// TIA Portal project "EdgeHowTos" (V16)

(* hardware
DEVICE "S71500/ET200MP station_1"  S7-1500 station
   slot 0: "Rail_0"  Rack  6ES7 590-1***0-0AA0
   slot 1: "PLC"  CPU 1513-1 PN  6ES7 513-1AL02-0AB0  V2.8
      slot 3: "CPU display_1"  6ES7591-1AA00-0AA0
      slot 32768: "PROFINET interface_1"  X1
         slot 32769: "Port_1"  X1 P1
         slot 32770: "Port_2"  X1 P2
      slot 34817: "Virtual CP interface port_1"  Virtual CP interface port  Virtual CP interface port
DEVICE "HMI"  TP900 Comfort
   slot 0: "HMI"  TP900 Comfort  6AV2 124-0JC01-0AX0  16.0.0.0
   slot 1: "HMI_RT_5"  TP900 Comfort  6AV2 124-0JC01-0AX0  16.0.0.0
   slot 5: "HMI._CP_1"  PROFINET Interface  16.0.0.0
      slot 1: "PROFINET Interface_1"  PROFINET Interface
         slot 1: "Port_1"  Port
         slot 2: "Port_2"  Port
   slot 7: "HMI.I/DP_CP_1"  MPI/DP Interface  16.0.0.0
*)

// ===== PLC "PLC"  CPU 1513-1 PN =====

VAR_GLOBAL   // PLC tag table "Default tag table"
   "Manipulator" AT %MW0 : Int;
END_VAR

VAR_GLOBAL CONSTANT   // PLC tag table "Default tag table"
   "STATE_FILL_TANK" : Int := 1;
   "STATE_HEAT_TANK" : Int := 2;
   "STATE_FILL_BOTTLE" : Int := 3;
   "STATE_SHIFT_BOTTLE" : Int := 4;
   "STATE_STOP" : Int := 5;
   "STATE_RESET" : Int := 6;
   "STATE_ERROR" : Int := 7;
   "ERROR_0_NO" : UInt := 0;
   "ERROR_1_CONNECTION" : UInt := 1;
   "ERROR_2_POWER" : UInt := 2;
   "ERROR_3_MANPOWER" : UInt := 3;
   "ERROR_4_CONVEYOR" : UInt := 4;
   "ERROR_5_VENTIL" : UInt := 5;
   "ERROR_6_HEATING" : UInt := 6;
   "ERROR_7_BOTTLE" : UInt := 7;
END_VAR

TYPE "typeHmi"
   STRUCT
      HMI_Start : Bool;   // trigger from hmi to start
      HMI_Stop : Bool;   // trigger from hmi to stop
      HMI_Reset : Bool;   // trigger from hmi to reset
      HMI_NextBottle : Bool;   // trigger from hmi to shift bottle
      HMI_Error : Bool;   // trigger from hmi to generate error
   END_STRUCT;
END_TYPE

TYPE "typeApp"
   STRUCT
      APP_Start : Bool;   // trigger from app to start
      APP_Stop : Bool;   // trigger from app to stop
      APP_Reset : Bool;   // trigger from app to reset
      APP_QRCode : String;   // string from app containing QR code (scanning app)
      APP_NextBottle : Bool;   // trigger from app to shift bottle
      APP_Error : Bool;   // trigger from app to generate error
      APP_Alarm : Bool;   // trigger from app to generate program alarm
   END_STRUCT;
END_TYPE

TYPE "typeSignals"
   STRUCT
      tankSignals : Struct
         actLevel : Real;   // actual level of tank [l]
         maxLevel : Bool;   // max level of tank reached
         actPressure : Real;   // actual pressure of tank [hPa]
         actTemperature : Real;   // actual temperature of tank [°C]
         maxTemperature : Bool;   // max level of temperature reached
      END_STRUCT;
      bottleSignals : Struct
         actLevel : Real;   // actual level of current bottle [l]
         maxLevel : Bool;   // max level of bottle reached
         outputTank : Real;   // Vout of Tank / Vin of bottle [m³/s]
      END_STRUCT;
      energySignals : Struct
         energyConsumptionFillingTank : Real;   // energy consumption during filling tank [Wh]
         waterConsumptionFillingTank : Real;   // water consumption during filling tank [l]
         energyConsumptionHeatingTank : Real;   // energy consumption during heating tank [Wh]
         energyConsumptionFillingBottles : Real;   // energy consumption during filling bottles [Wh]
         gasConsumptionHeatingTank : Real;   // gas consumption during heating tank [Wh]
      END_STRUCT;
      alarm : Word;   // alarm bit
   END_STRUCT;
END_TYPE

TYPE "typeOperate"
   STRUCT
      extModeActive : Bool := false;   // true = activate external model / simulation
      state : "typeState";   // operating state
      machineState : Int := 0;   // see user constants (1 = filling tank, 2 = heating tank, 3 = filling bottle, 4 = shifting bottle, 5 = stop, 6 = reset)
   END_STRUCT;
END_TYPE

TYPE "typeModel"
   STRUCT
      cycleTime : Real;   // cycle time[s]
      tank : Struct   // model struct of tank
         AT : Real;   // surface area of tank [m²]
         H : Real;   // high of tank [m]
         Vin : Real;   // incoming volume flow [l/min]
         maxLevel : Real;   // max level of tank [m³]
         roomTemperature : Real;   // room temperature of tank [°C]
         maxTemperature : Real;   // max temperature of tank [°C]
         density : Real;   // liquid density [kg/m³]
      END_STRUCT;
      bottle : Struct   // model struct of bottle
         maxLevel : Real;   // max level of bottle [m³]
         AB : Real;   // surface area of filling hole to fill bottle [m²]
      END_STRUCT;
   END_STRUCT;
END_TYPE

TYPE "typeProcess"
   STRUCT
      productId : UDInt;   // product id of current bottle
      numberProduced : UDInt;   // number of filled bottles
      numberFaulty : UDInt;   // number of faulty bottles
      batchId : UDInt;   // batch id (according to tank filling)
   END_STRUCT;
END_TYPE

TYPE "typeState"
   STRUCT
      FillingTank : Bool;   // filling tank
      HeatingTank : Bool;   // heating tank
      FillingBottle : Bool;   // filling bottle
      ShiftingBottle : Bool;   // shifting bottle
      Stop : Bool;   // stop filling application
      Reset : Bool;   // reset application
      Error : Bool;   // error within filling application
   END_STRUCT;
END_TYPE

TYPE "typeInfo"
   STRUCT
      "version" : String;   // current version of the project
      "date" : String;   // last change date of the project
   END_STRUCT;
END_TYPE

TYPE "typeError"
   STRUCT
      errorSimulation : Bool := true;   // activate simulation
      errorTrigger : Bool := false;   // trigger manual error simulation
      errorDuration : Time := T#120s;   // error duration for simlation
      errorCode : UInt := 0;   // error code for error analysis
   END_STRUCT;
END_TYPE

DATA_BLOCK "GDB"   // DB1
{ S7_Optimized_Access := 'FALSE' }
VERSION : 0.1
   VAR
      operate : "typeOperate";   // application operation
      model : "typeModel";   // model parameter
      externalSignals : "typeSignals";   // signals from external model
      signals : "typeSignals";   // current signals from tank and bottle
      process : "typeProcess";   // current process information
      hmiSignals : "typeHmi";   // signals from hmi
      appSignals : "typeApp";   // signals from edge app
      projectInfo : "typeInfo";   // infos regarding this TIA project
      errors : "typeError";
   END_VAR
BEGIN
   model.tank.H := 2.0;
   model.tank.AT := 0.8;
   operate.extModeActive := false;
   model.tank.maxTemperature := 80.0;
   model.tank.maxLevel := 1.6;
   model.bottle.maxLevel := 0.1;
   model.cycleTime := 0.01;
   model.tank.roomTemperature := 20.0;
   model.tank.Vin := 500.0;
   model.bottle.AB := 0.001;
   process.productId := 0;
   process.numberProduced := 0;
   process.numberFaulty := 0;
   model.tank.density := 997.0;
   hmiSignals.HMI_Start := true;
   projectInfo."version" := 'V1.1';
   projectInfo."date" := '2024-04-18';
END_DATA_BLOCK

DATA_BLOCK "DB_1_Sequence"   // DB2
{ S7_Optimized_Access := 'TRUE' }
VERSION : 0.1
// stored: InstanceOfName FB_1_Sequence
"FB_1_Sequence"
BEGIN
END_DATA_BLOCK

DATA_BLOCK "DB_2_Filling_DB"   // DB3
{ S7_Optimized_Access := 'TRUE' }
VERSION : 0.1
// stored: InstanceOfName FB_2_Filling
"FB_2_Filling"
BEGIN
END_DATA_BLOCK

DATA_BLOCK "DB_3_Simulation"   // DB4
{ S7_Optimized_Access := 'TRUE' }
VERSION : 0.1
// stored: InstanceOfName FB_3_Simulation
"FB_3_Simulation"
BEGIN
END_DATA_BLOCK

FUNCTION_BLOCK "FB_1_Sequence"   // FB2, FBD
{ S7_Optimized_Access := 'TRUE' }
VERSION : 0.1
   VAR_INPUT
      model : "typeModel";   // model parameter
      externalSignals : "typeSignals";   // signals from external model
   END_VAR
   VAR_IN_OUT
      operate : "typeOperate";   // application operation
      signals : "typeSignals";   // current signals from tank
      process : "typeProcess";   // current process information
      hmi : "typeHmi";   // signals from hmi
      app : "typeApp";   // signals from app
      errors : "typeError";
   END_VAR
   VAR
      statStart : Bool;   // trigger for start command
      statStop : Bool;   // trigger for stop command
      statReset : Bool;   // trigger for reset command
      statInit : Bool := true;   // helper variable to initialize some parameters
      statNextBottle : Bool;   // trigger to shift next bottle
      statError : Bool;   // trigger to set error
      statState : Int;   // memory for reactivating state after STOP
      statAlarm : Bool;   // trigger to generate program alarm
      statMemoryStart : Bool;
      statMemoryStop : Bool;
      statMemoryReset : Bool;
      statMemoryNextBottle : Bool;
      statMemoryError : Bool;
      statHmiStateStart : Bool;   // helper for hmi (true, if state 1-4)
      statShiftingTimer : Int;
      statShiftingTimerTrigger : Bool;
      statShiftingTrigger : Bool;
      statShiftingTimerDone : Bool;
      statHmiQrCodeReceived : Bool;
      statHMIQrCodeReceivedTrigger : Bool;
      statQrCodeTrigger : Bool;
      statTankEmpty : Bool;   // trigger when tank is empty
      statTankEmptyMemory : Bool;   // tank empty memory
      statOverflow : Bool;   // overflow of counter "numberProduced"
      statOverflowStartTrigger : Bool;   // trigger to start after overflow
      statOverflowStartMemory : Bool;
      Program_Alarm : Program_Alarm;
   END_VAR
   VAR_TEMP
      tempQrCodeLen : Int;
      tempProgramAlarmError : Bool;
      tempProgramAlarmStatus : Word;
      tempAlarmStateError : Bool;
      tempAlarmStateStatus : Word;
   END_VAR
   VAR_TEMP   // added for the SCL form of the ladder/FBD networks
      _w1 : Bool;
      _w2 : Bool;
      _w3 : Bool;
      _w4 : Bool;
   END_VAR
BEGIN

REGION Network 1: Handling signals from hmi or app
   // --[P]-- (positive signal edge) -> stat-Variable becomes true for one cycle
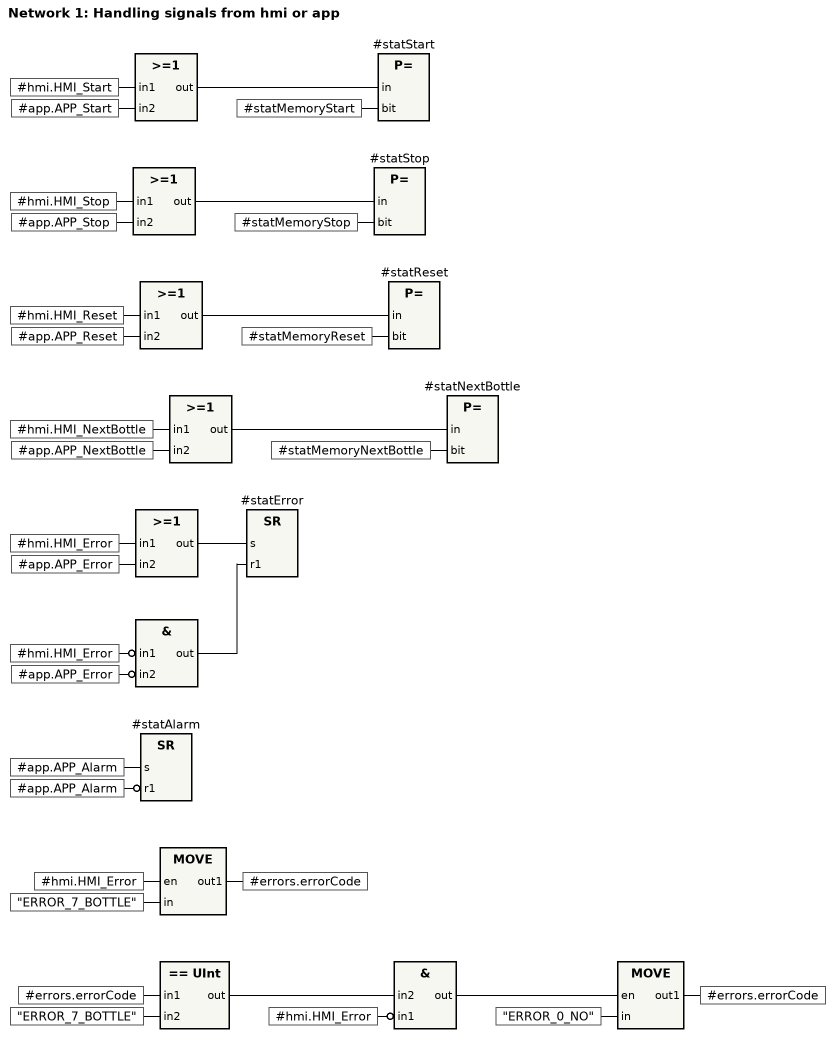
   #_w1 := #hmi.HMI_Start OR #app.APP_Start;
   #statStart := #_w1 AND NOT #statMemoryStart;   // rising edge
   #statMemoryStart := #_w1;
   #_w2 := #hmi.HMI_Stop OR #app.APP_Stop;
   #statStop := #_w2 AND NOT #statMemoryStop;   // rising edge
   #statMemoryStop := #_w2;
   #_w3 := #hmi.HMI_Reset OR #app.APP_Reset;
   #statReset := #_w3 AND NOT #statMemoryReset;   // rising edge
   #statMemoryReset := #_w3;
   #_w4 := #hmi.HMI_NextBottle OR #app.APP_NextBottle;
   #statNextBottle := #_w4 AND NOT #statMemoryNextBottle;   // rising edge
   #statMemoryNextBottle := #_w4;
   IF #hmi.HMI_Error OR #app.APP_Error THEN
       #statError := TRUE;   // SR flip-flop
   END_IF;
   IF NOT #hmi.HMI_Error AND NOT #app.APP_Error THEN #statError := FALSE; END_IF;
   IF #app.APP_Alarm THEN
       #statAlarm := TRUE;   // SR flip-flop
   END_IF;
   IF NOT #app.APP_Alarm THEN #statAlarm := FALSE; END_IF;
   IF #hmi.HMI_Error THEN #errors.errorCode := "ERROR_7_BOTTLE"; END_IF;
   IF (#errors.errorCode = "ERROR_7_BOTTLE") AND NOT #hmi.HMI_Error THEN
       #errors.errorCode := "ERROR_0_NO";
   END_IF;
END_REGION

REGION Network 2: Reset signals from hmi or app
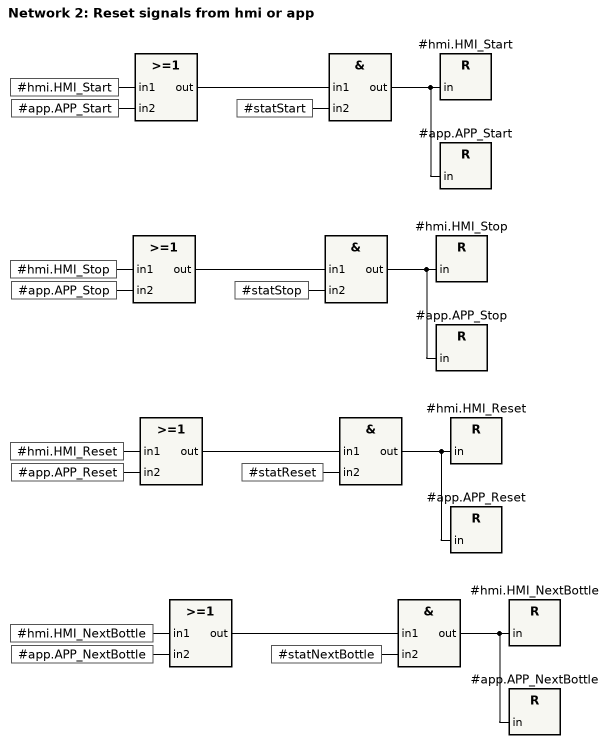
   #_w1 := (#hmi.HMI_Start OR #app.APP_Start) AND #statStart;
   IF #_w1 THEN
       #hmi.HMI_Start := FALSE;
       #app.APP_Start := FALSE;
   END_IF;
   #_w2 := (#hmi.HMI_Stop OR #app.APP_Stop) AND #statStop;
   IF #_w2 THEN
       #hmi.HMI_Stop := FALSE;
       #app.APP_Stop := FALSE;
   END_IF;
   #_w3 := (#hmi.HMI_Reset OR #app.APP_Reset) AND #statReset;
   IF #_w3 THEN
       #hmi.HMI_Reset := FALSE;
       #app.APP_Reset := FALSE;
   END_IF;
   #_w4 := (#hmi.HMI_NextBottle OR #app.APP_NextBottle) AND #statNextBottle;
   IF #_w4 THEN
       #hmi.HMI_NextBottle := FALSE;
       #app.APP_NextBottle := FALSE;
   END_IF;
END_REGION

REGION Network 3: Helper for hmi display
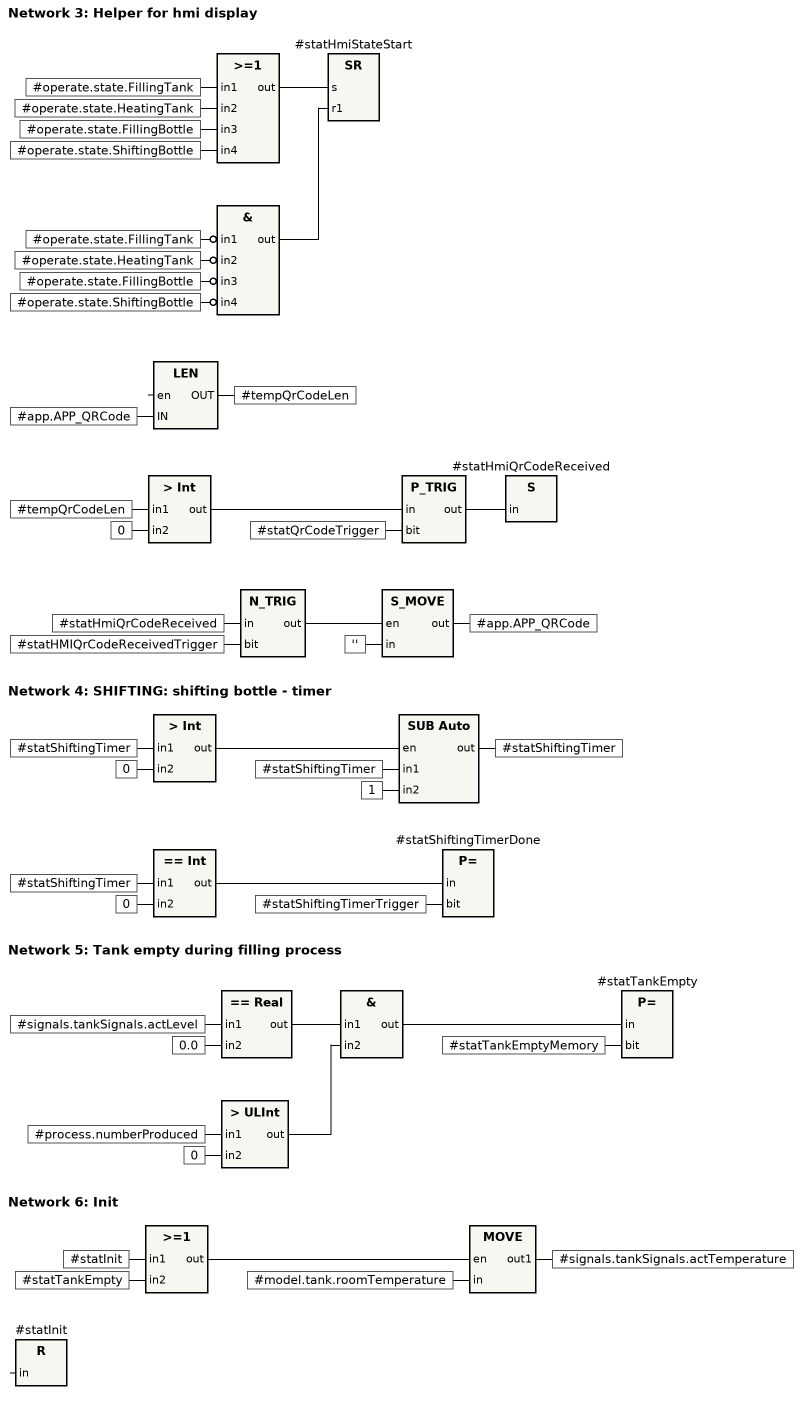
   IF #operate.state.FillingTank OR #operate.state.HeatingTank OR #operate.state.FillingBottle OR #operate.state.ShiftingBottle THEN
       #statHmiStateStart := TRUE;   // SR flip-flop
   END_IF;
   IF NOT #operate.state.FillingTank AND NOT #operate.state.HeatingTank AND NOT #operate.state.FillingBottle AND NOT #operate.state.ShiftingBottle THEN
       #statHmiStateStart := FALSE;
   END_IF;
   #tempQrCodeLen := LEN(IN := #app.APP_QRCode);
   #_w1 := #tempQrCodeLen > 0;
   #_w2 := #_w1 AND NOT #statQrCodeTrigger;   // rising edge
   #statQrCodeTrigger := #_w1;
   IF #_w2 THEN #statHmiQrCodeReceived := TRUE; END_IF;
   #_w3 := NOT #statHmiQrCodeReceived AND #statHMIQrCodeReceivedTrigger;   // falling edge
   #statHMIQrCodeReceivedTrigger := #statHmiQrCodeReceived;
   IF #_w3 THEN #app.APP_QRCode := ''; END_IF;
END_REGION

REGION Network 4: SHIFTING: shifting bottle - timer
   IF #statShiftingTimer > 0 THEN #statShiftingTimer := #statShiftingTimer - 1; END_IF;
   #_w1 := #statShiftingTimer = 0;
   #statShiftingTimerDone := #_w1 AND NOT #statShiftingTimerTrigger;   // rising edge
   #statShiftingTimerTrigger := #_w1;
END_REGION

REGION Network 5: Tank empty during filling process
   #_w1 := (#signals.tankSignals.actLevel = 0.0) AND (#process.numberProduced > 0);
   #statTankEmpty := #_w1 AND NOT #statTankEmptyMemory;   // rising edge
   #statTankEmptyMemory := #_w1;
END_REGION

REGION Network 6: Init
   IF #statInit OR #statTankEmpty THEN
       #signals.tankSignals.actTemperature := #model.tank.roomTemperature;
   END_IF;
   #statInit := FALSE;
END_REGION

REGION Network 7: Filling tank
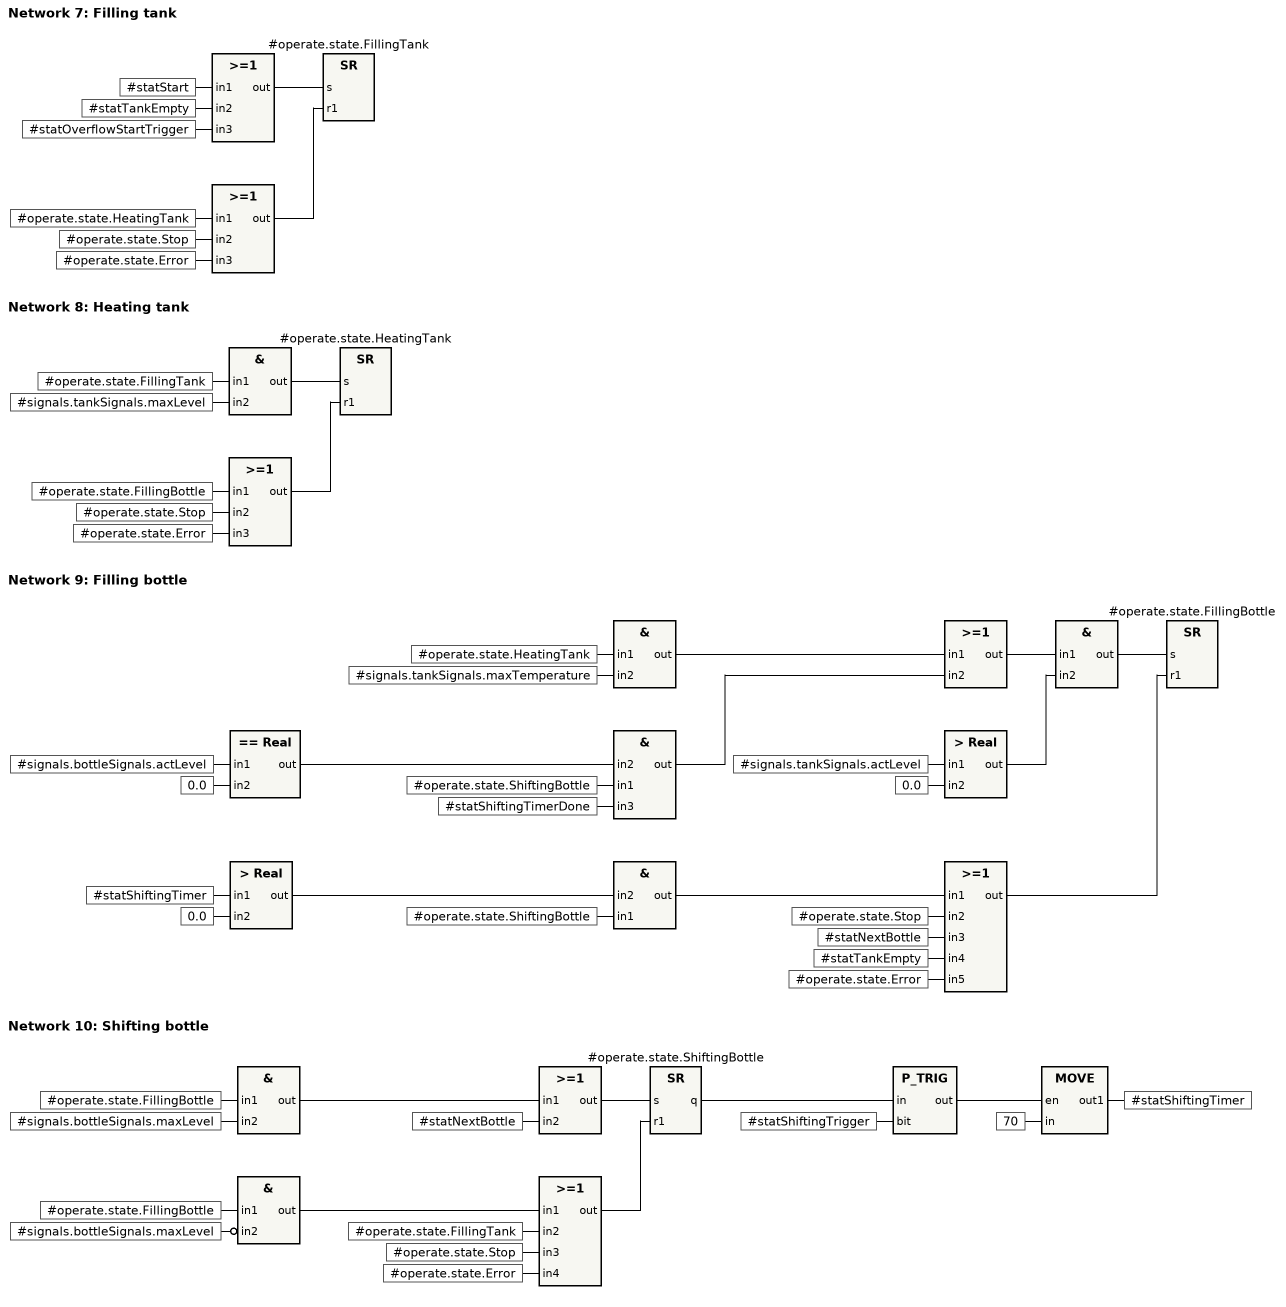
   IF #statStart OR #statTankEmpty OR #statOverflowStartTrigger THEN
       #operate.state.FillingTank := TRUE;   // SR flip-flop
   END_IF;
   IF #operate.state.HeatingTank OR #operate.state.Stop OR #operate.state.Error THEN
       #operate.state.FillingTank := FALSE;
   END_IF;
END_REGION

REGION Network 8: Heating tank
   IF #operate.state.FillingTank AND #signals.tankSignals.maxLevel THEN
       #operate.state.HeatingTank := TRUE;   // SR flip-flop
   END_IF;
   IF #operate.state.FillingBottle OR #operate.state.Stop OR #operate.state.Error THEN
       #operate.state.HeatingTank := FALSE;
   END_IF;
END_REGION

REGION Network 9: Filling bottle
   IF ((#operate.state.HeatingTank AND #signals.tankSignals.maxTemperature) OR ((#signals.bottleSignals.actLevel = 0.0) AND #operate.state.ShiftingBottle AND #statShiftingTimerDone)) AND (#signals.tankSignals.actLevel > 0.0) THEN
       #operate.state.FillingBottle := TRUE;   // SR flip-flop
   END_IF;
   IF ((#statShiftingTimer > 0.0) AND #operate.state.ShiftingBottle) OR #operate.state.Stop OR #statNextBottle OR #statTankEmpty OR #operate.state.Error THEN
       #operate.state.FillingBottle := FALSE;
   END_IF;
END_REGION

REGION Network 10: Shifting bottle
   IF (#operate.state.FillingBottle AND #signals.bottleSignals.maxLevel) OR #statNextBottle THEN
       #operate.state.ShiftingBottle := TRUE;   // SR flip-flop
   END_IF;
   IF (#operate.state.FillingBottle AND NOT #signals.bottleSignals.maxLevel) OR #operate.state.FillingTank OR #operate.state.Stop OR #operate.state.Error THEN
       #operate.state.ShiftingBottle := FALSE;
   END_IF;
   #_w1 := #operate.state.ShiftingBottle AND NOT #statShiftingTrigger;   // rising edge
   #statShiftingTrigger := #operate.state.ShiftingBottle;
   IF #_w1 THEN #statShiftingTimer := 70; END_IF;
END_REGION

REGION Network 11: Catch overflow
   // If max of UDINT is reached
   // > Stop (automatically)
   // > Reset (automatically)
   // > Start (automatically)
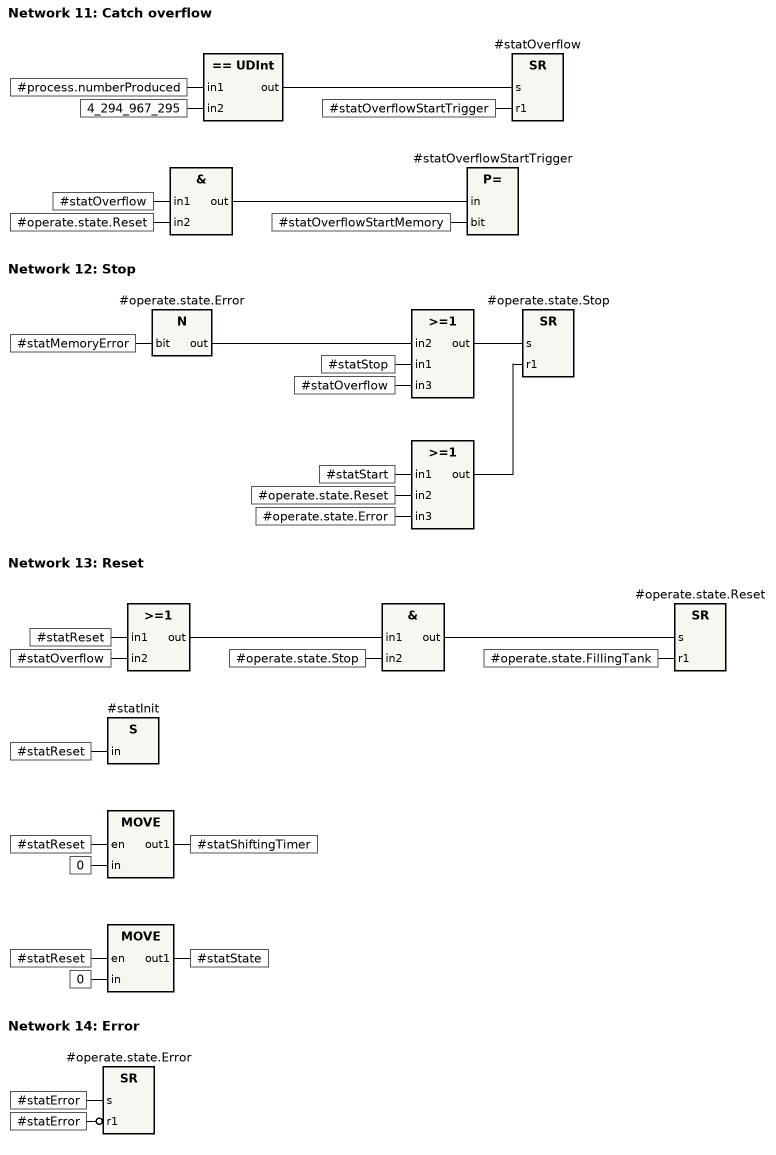
   IF #process.numberProduced = 4_294_967_295 THEN
       #statOverflow := TRUE;   // SR flip-flop
   END_IF;
   IF #statOverflowStartTrigger THEN #statOverflow := FALSE; END_IF;
   #_w1 := #statOverflow AND #operate.state.Reset;
   #statOverflowStartTrigger := #_w1 AND NOT #statOverflowStartMemory;   // rising edge
   #statOverflowStartMemory := #_w1;
END_REGION

REGION Network 12: Stop
   #_w1 := NOT #operate.state.Error AND #statMemoryError;   // falling edge of #operate.state.Error
   #statMemoryError := #operate.state.Error;
   IF #_w1 OR #statStop OR #statOverflow THEN
       #operate.state.Stop := TRUE;   // SR flip-flop
   END_IF;
   IF #statStart OR #operate.state.Reset OR #operate.state.Error THEN #operate.state.Stop := FALSE; END_IF;
END_REGION

REGION Network 13: Reset
   IF (#statReset OR #statOverflow) AND #operate.state.Stop THEN
       #operate.state.Reset := TRUE;   // SR flip-flop
   END_IF;
   IF #operate.state.FillingTank THEN #operate.state.Reset := FALSE; END_IF;
   IF #statReset THEN
       #statInit := TRUE;
       #statShiftingTimer := 0;
       #statState := 0;
   END_IF;
END_REGION

REGION Network 14: Error
   IF #statError THEN
       #operate.state.Error := TRUE;   // SR flip-flop
   END_IF;
   IF NOT #statError THEN #operate.state.Error := FALSE; END_IF;
END_REGION

REGION Network 15: Set machine state
   // 1 = filling tank
   // 2 = heating tank
   // 3 = filling bottle
   // 4 = shifting bottle
   // 5 = stop
   // 6 = reset
   // 7 = error
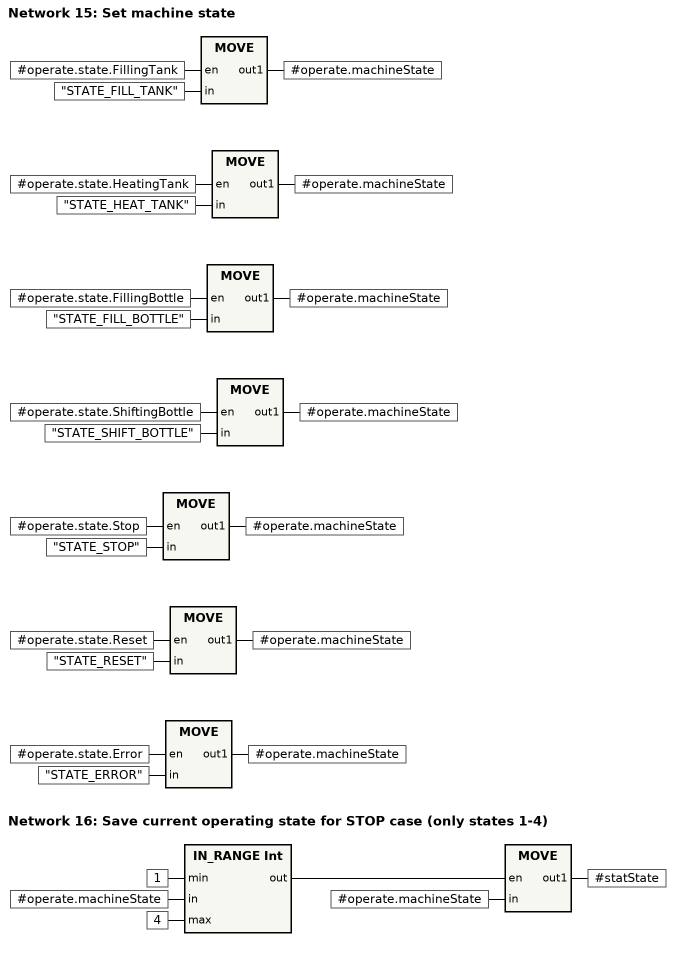
   IF #operate.state.FillingTank THEN #operate.machineState := "STATE_FILL_TANK"; END_IF;
   IF #operate.state.HeatingTank THEN #operate.machineState := "STATE_HEAT_TANK"; END_IF;
   IF #operate.state.FillingBottle THEN #operate.machineState := "STATE_FILL_BOTTLE"; END_IF;
   IF #operate.state.ShiftingBottle THEN #operate.machineState := "STATE_SHIFT_BOTTLE"; END_IF;
   IF #operate.state.Stop THEN #operate.machineState := "STATE_STOP"; END_IF;
   IF #operate.state.Reset THEN #operate.machineState := "STATE_RESET"; END_IF;
   IF #operate.state.Error THEN #operate.machineState := "STATE_ERROR"; END_IF;
END_REGION

REGION Network 16: Save current operating state for STOP case (only states 1-4)
   // 1 = filling tank
   // 2 = heating tank
   // 3 = filling bottle
   // 4 = shifting bottle
   IF (1 <= #operate.machineState) AND (#operate.machineState <= 4) THEN
       #statState := #operate.machineState;
   END_IF;
END_REGION

REGION Network 17: Reactivate old state after STOP
   // 1 = filling tank
   // 2 = heating tank
   // 3 = filling bottle
   // 4 = shifting bottle
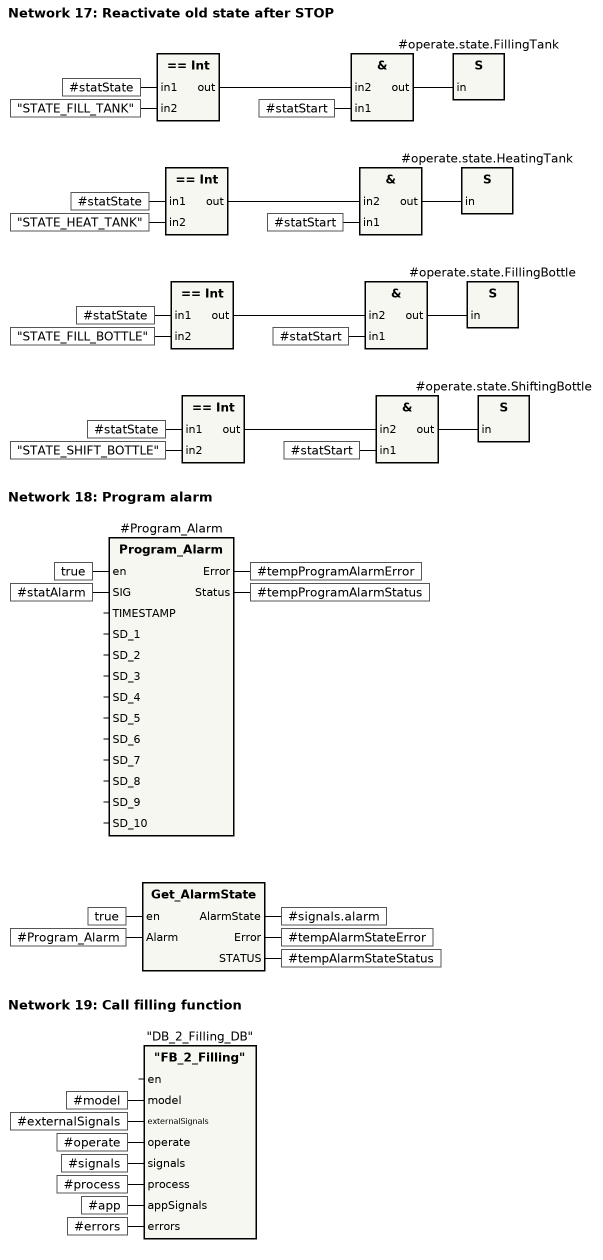
   IF (#statState = "STATE_FILL_TANK") AND #statStart THEN #operate.state.FillingTank := TRUE; END_IF;
   IF (#statState = "STATE_HEAT_TANK") AND #statStart THEN #operate.state.HeatingTank := TRUE; END_IF;
   IF (#statState = "STATE_FILL_BOTTLE") AND #statStart THEN #operate.state.FillingBottle := TRUE; END_IF;
   IF (#statState = "STATE_SHIFT_BOTTLE") AND #statStart THEN #operate.state.ShiftingBottle := TRUE; END_IF;
END_REGION

REGION Network 18: Program alarm
   // no SCL statement known for Get_AlarmState: written as a call
   IF true THEN
       #Program_Alarm(SIG := #statAlarm, Error => #tempProgramAlarmError, Status => #tempProgramAlarmStatus);   // Program_Alarm
       Get_AlarmState(Alarm := #Program_Alarm,
                      AlarmState => #signals.alarm,
                      Error => #tempAlarmStateError,
                      STATUS => #tempAlarmStateStatus);
   END_IF;
END_REGION

REGION Network 19: Call filling function
   "DB_2_Filling_DB"(model := #model,   // "FB_2_Filling"
                     externalSignals := #externalSignals,
                     operate := #operate,
                     signals := #signals,
                     process := #process,
                     appSignals := #app,
                     errors := #errors);
END_REGION
END_FUNCTION_BLOCK

FUNCTION_BLOCK "FB_2_Filling"   // FB3, FBD
TITLE = Filling process
{ S7_Optimized_Access := 'TRUE' }
VERSION : 0.1
   VAR_INPUT
      model : "typeModel";   // model parameter
      externalSignals : "typeSignals";   // signals from external model
   END_VAR
   VAR_IN_OUT
      operate : "typeOperate";   // application operation
      signals : "typeSignals";   // current signals from tank
      process : "typeProcess";   // current process information
      appSignals : "typeApp";
      errors : "typeError";   // error information
   END_VAR
   VAR
      statShiftingBottle : Bool;
      statShiftingTrigger : Bool;
      statShiftingTimer : Int;
      statHmiBottleLevel : Real;   // parameter for HMI to show current bottle level
      statHmiDoShift : Bool;   // trigger for HMI to shift bottles
      statHmiFaultyBottle : Bool;   // trigger for HMI for faulty bottle
      statFillingTankTrigger : Bool;
   END_VAR
   VAR_TEMP
      tempBottleMaxLevel : Real;
   END_VAR
   VAR_TEMP   // added for the SCL form of the ladder/FBD networks
      _w1 : Bool;
      _w2 : Bool;
   END_VAR
BEGIN

REGION Network 1: Calculation of params
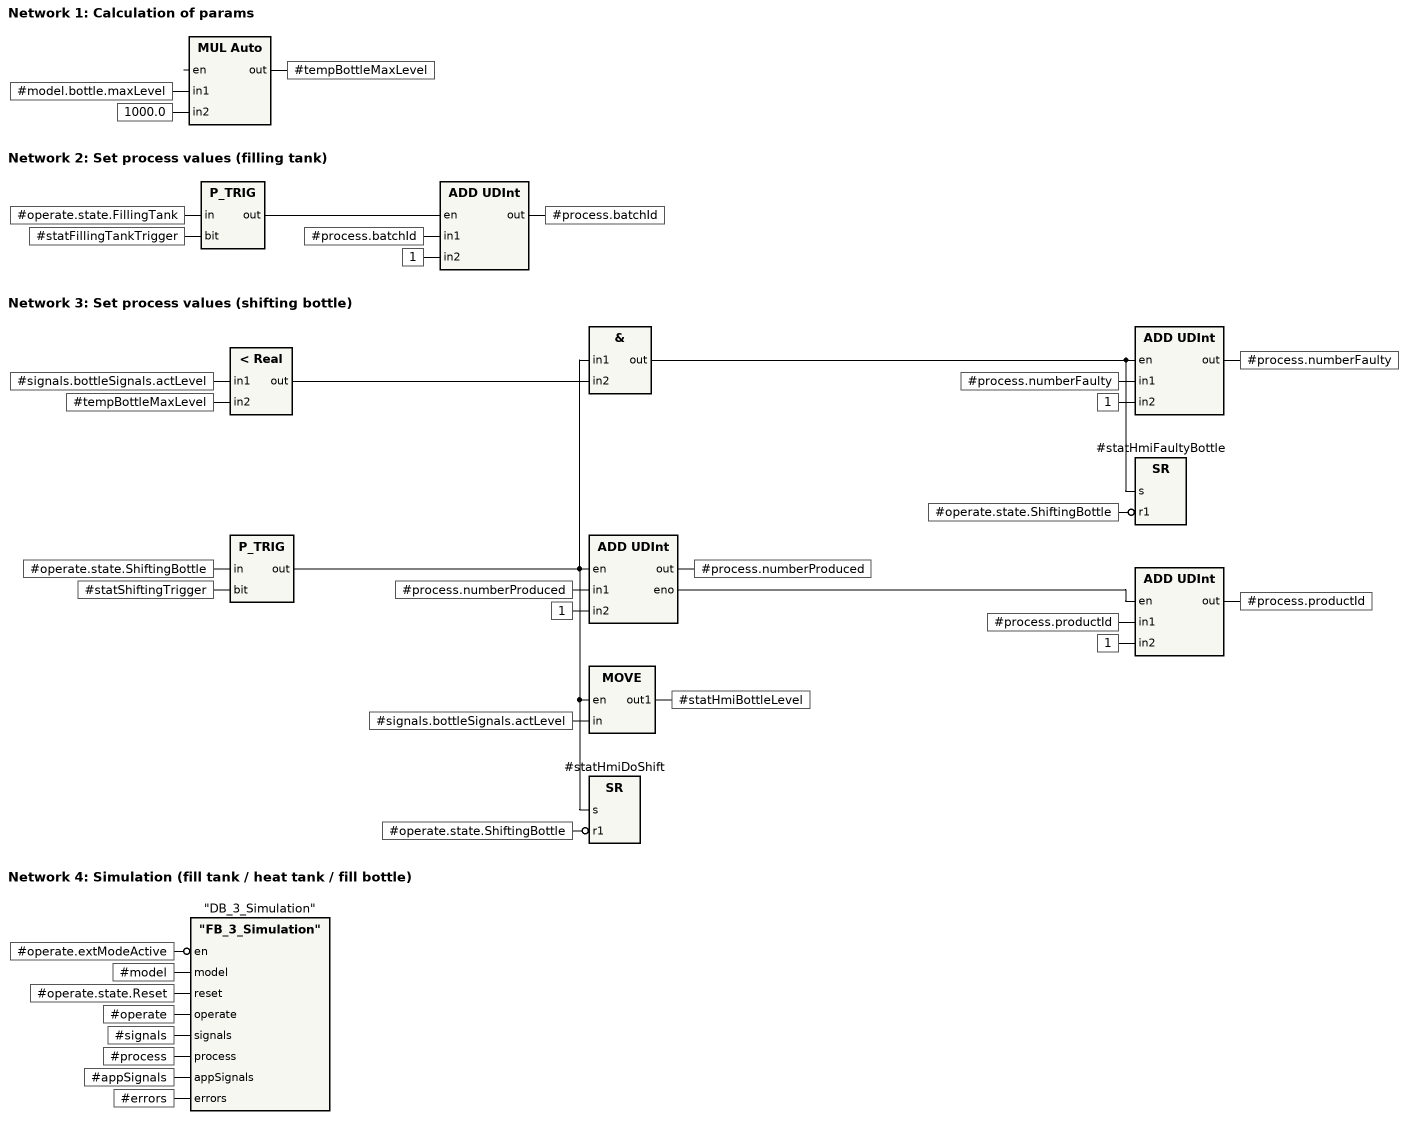
   #tempBottleMaxLevel := #model.bottle.maxLevel * 1000.0;
END_REGION

REGION Network 2: Set process values (filling tank)
   #_w1 := #operate.state.FillingTank AND NOT #statFillingTankTrigger;   // rising edge
   #statFillingTankTrigger := #operate.state.FillingTank;
   IF #_w1 THEN #process.batchId := #process.batchId + 1; END_IF;
END_REGION

REGION Network 3: Set process values (shifting bottle)
   #_w1 := #operate.state.ShiftingBottle AND NOT #statShiftingTrigger;   // rising edge
   #statShiftingTrigger := #operate.state.ShiftingBottle;
   IF #_w1 THEN
       #process.numberProduced := #process.numberProduced + 1;
       #process.productId := #process.productId + 1;
   END_IF;
   #_w2 := #_w1 AND (#signals.bottleSignals.actLevel < #tempBottleMaxLevel);
   IF #_w2 THEN
       #process.numberFaulty := #process.numberFaulty + 1;
       #statHmiFaultyBottle := TRUE;   // SR flip-flop
   END_IF;
   IF NOT #operate.state.ShiftingBottle THEN #statHmiFaultyBottle := FALSE; END_IF;
   IF #_w1 THEN
       #statHmiBottleLevel := #signals.bottleSignals.actLevel;
       #statHmiDoShift := TRUE;   // SR flip-flop
   END_IF;
   IF NOT #operate.state.ShiftingBottle THEN #statHmiDoShift := FALSE; END_IF;
END_REGION

REGION Network 4: Simulation (fill tank / heat tank / fill bottle)
   IF NOT #operate.extModeActive THEN
       "DB_3_Simulation"(model := #model,   // "FB_3_Simulation"
                         reset := #operate.state.Reset,
                         operate := #operate,
                         signals := #signals,
                         process := #process,
                         appSignals := #appSignals,
                         errors := #errors);
   END_IF;
END_REGION

REGION Network 5: Reset process parameter
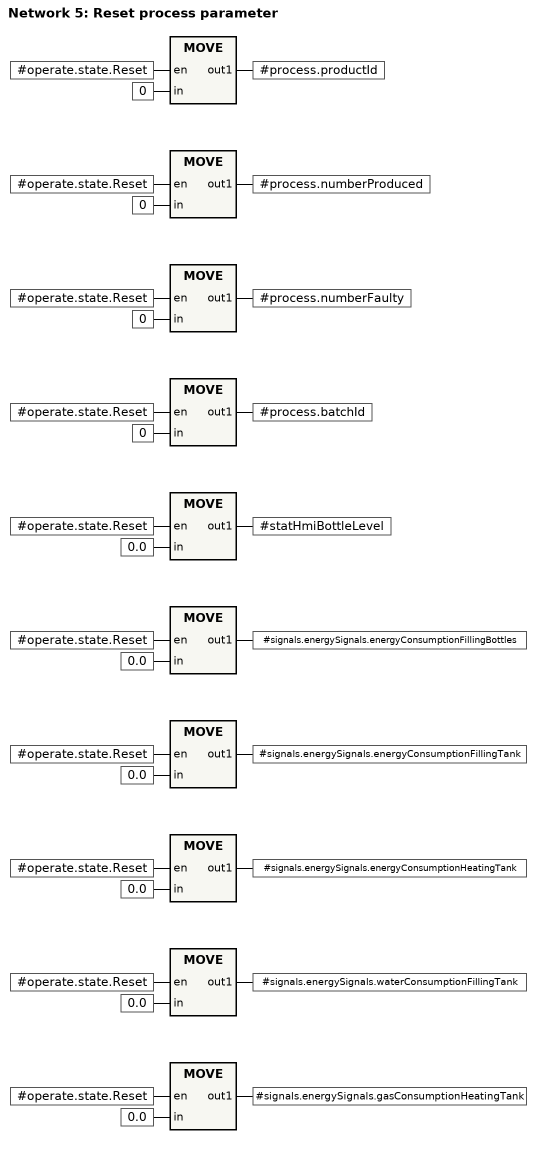
   IF #operate.state.Reset THEN
       #process.productId := 0;
       #process.numberProduced := 0;
       #process.numberFaulty := 0;
       #process.batchId := 0;
       #statHmiBottleLevel := 0.0;
       #signals.energySignals.energyConsumptionFillingBottles := 0.0;
       #signals.energySignals.energyConsumptionFillingTank := 0.0;
       #signals.energySignals.energyConsumptionHeatingTank := 0.0;
       #signals.energySignals.waterConsumptionFillingTank := 0.0;
       #signals.energySignals.gasConsumptionHeatingTank := 0.0;
   END_IF;
END_REGION
END_FUNCTION_BLOCK

FUNCTION_BLOCK "FB_3_Simulation"   // FB4, FBD
TITLE = Model Tank Level
{ S7_Optimized_Access := 'TRUE' }
VERSION : 0.1
   VAR_INPUT
      model : "typeModel";   // model parameter
      reset : Bool;   // reset tanklevel
      operate : "typeOperate";   // operate parameter
   END_VAR
   VAR_IN_OUT
      signals : "typeSignals";   // current signals from tank
      process : "typeProcess";   // current process parameters
      appSignals : "typeApp";
      errors : "typeError";
   END_VAR
   VAR
      "statVinl/min" : Real;   // Vin[l/min]
      "statVinM3/S" : Real;   // Vin [m³/s]
      statInputTanklevel : Real;   // TANK: input tank level for LSim_I [m³]
      statTankLevelSqrt : Real;   // TANK: sqrt of tank level [m³]
      statOutGainSqrt : Real;   // TANK: sqrt of GAIN_SQRT
      statOutGainDiv : Real;   // TANK: divide AB/AT
      statOutGainValue : Real;   // TANK: output gain value
      statVoutSwitch : Real;   // TANK: Vout switch
      statVoutMultiplier : Real;   // TANK: tank level sqrt *output gain value [m³]
      statTankLevel : Real;   // TANK: current level of tank (m³)
      statLiquidMass : Real;   // TANK: liquid mass [kg]
      statLiquidPower : Real;   // TANK: liquid power [N]
      statLiquidPressure_Pa : Real;   // TANK: liquid pressure [Pa]
      instLSim_I_tank : "LSim_I";   // TANK: instance of LSim_I
      statPT1in1 : Real;   // HEAT: input PT1_1
      statPT1out1 : Real;   // HEAT: output PT1_1
      statPT1out2 : Real;   // HEAT: output PT1_2
      instLSim_PT1_1 : "LSim_PT1";   // HEAT: instance PT1 1
      instLSim_PT1_2 : "LSim_PT1";   // HEAT: instance PT1 2
      instLSim_PT1_3 : "LSim_PT1";   // HEAT: instance PT1 3
      instLSim_PT3 : "LSim_PT3";   // HEAT: instance of PT3
      statPT3in : Real;   // HEAT: input value for PT3
      instLSim_I_bottle : "LSim_I";   // BOTTLE: instance of LSim_I
      statBottleLevel : Real;   // BOTTLE: Input bottle level for LSim_I
      statHeatTmLag : Real;   // HEAT: parameter for tmLag1
      statResetHeatingTrigger : Bool;   // trigger for resetting heating
      statResetHeatingMem : Bool;
      statHeatingActive : Bool;   // is set, when heating is active (to 80°C)
      statTriggerResetEnergy : Bool;
      statStopMem : Bool;   // trigger memory for stop
      statShiftingMem : Bool;   // trigger memory for shifting bottle
      statErrorMem : Bool;   // trigger memory for new error
      statResetError : Bool;   // helper bit for error > start workflow
      instTimerError : IEC_TIMER;
      statStart : Bool;   // helper to go in Start state
   END_VAR
   VAR_TEMP
      tempValue : Real;
      tempEnableHeating : Bool;   // enable heating controller
      tempRandomNumber : Real;
      tempRandomNumber1 : Real;
      tempRandomNumber2 : Real;
      tempRandomNumber3 : Int;   // random number for faulty bottle generation
      tempRandomNumber4 : UInt;   // random number for error code
      tempRandomNumber5 : UInt;   // random number for error state
      tempStopTrigger : Bool;   // trigger for stop
      tempShiftingTrigger : Bool;   // trigger for shifting bottle
      tempErrorTrigger : Bool;   // trigger for new error
   END_VAR
   VAR CONSTANT
      RECALC_VIN : Real := 1.667E-05;   // TANK: 1.667E-05 (1/1000 * 1/60), recalc Vin l/min -> m³/s
      GAIN_SQRT : Real := 19.62;   // TANK: 2*9.81
      GAIN : Real := 1.0;   // HEAT: gain value
      ACCELERATION : Real := 9.81;   // gravitational acceleration (a = 9,81 m/s²)
   END_VAR
   VAR_TEMP   // added for the SCL form of the ladder/FBD networks
      _w1 : Bool;
   END_VAR
BEGIN

REGION Network 1: TANK: Vin switch [l/min]
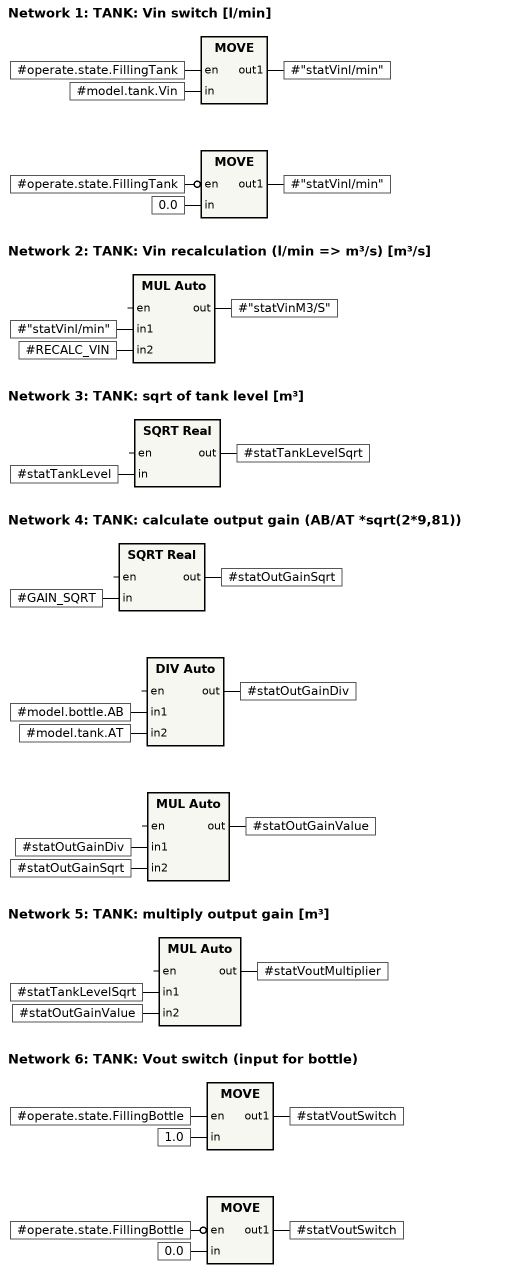
   IF #operate.state.FillingTank THEN #"statVinl/min" := #model.tank.Vin; END_IF;
   IF NOT #operate.state.FillingTank THEN #"statVinl/min" := 0.0; END_IF;
END_REGION

REGION Network 2: TANK: Vin recalculation (l/min => m³/s) [m³/s]
   #"statVinM3/S" := #"statVinl/min" * #RECALC_VIN;
END_REGION

REGION Network 3: TANK: sqrt of tank level [m³]
   #statTankLevelSqrt := SQRT(#statTankLevel);
END_REGION

REGION Network 4: TANK: calculate output gain (AB/AT *sqrt(2*9,81))
   #statOutGainSqrt := SQRT(#GAIN_SQRT);
   #statOutGainDiv := #model.bottle.AB / #model.tank.AT;
   #statOutGainValue := #statOutGainDiv * #statOutGainSqrt;
END_REGION

REGION Network 5: TANK: multiply output gain [m³]
   #statVoutMultiplier := #statTankLevelSqrt * #statOutGainValue;
END_REGION

REGION Network 6: TANK: Vout switch (input for bottle)
   IF #operate.state.FillingBottle THEN #statVoutSwitch := 1.0; END_IF;
   IF NOT #operate.state.FillingBottle THEN #statVoutSwitch := 0.0; END_IF;
END_REGION

REGION Network 7: TANK: Vout multiplier [m³/s]
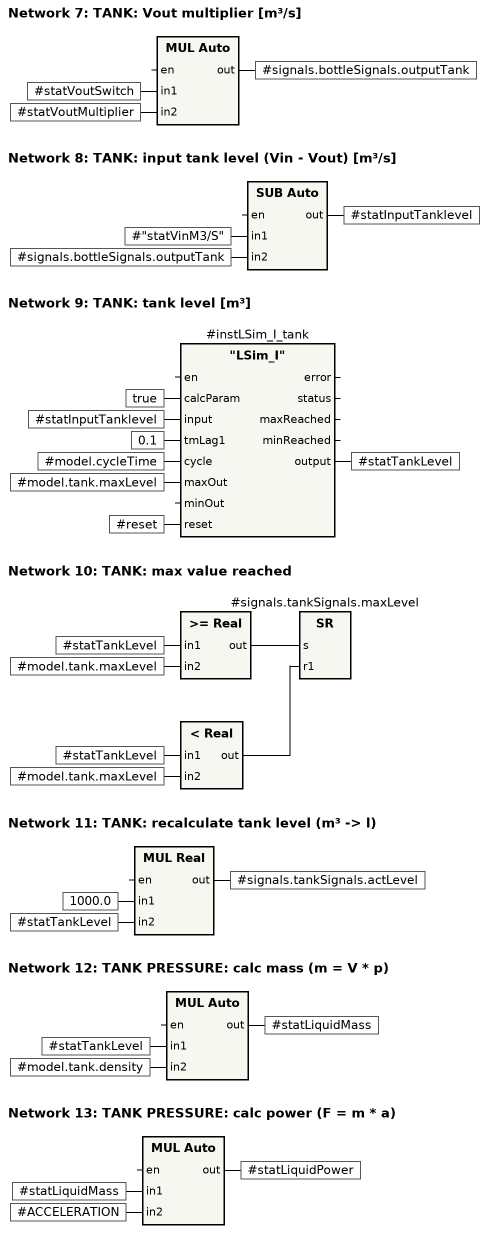
   #signals.bottleSignals.outputTank := #statVoutSwitch * #statVoutMultiplier;
END_REGION

REGION Network 8: TANK: input tank level (Vin - Vout) [m³/s]
   #statInputTanklevel := #"statVinM3/S" - #signals.bottleSignals.outputTank;
END_REGION

REGION Network 9: TANK: tank level [m³]
   #instLSim_I_tank(calcParam := true,   // "LSim_I"
                    input := #statInputTanklevel,
                    tmLag1 := 0.1,
                    cycle := #model.cycleTime,
                    maxOut := #model.tank.maxLevel,
                    reset := #reset,
                    output => #statTankLevel);
END_REGION

REGION Network 10: TANK: max value reached
   IF #statTankLevel >= #model.tank.maxLevel THEN
       #signals.tankSignals.maxLevel := TRUE;   // SR flip-flop
   END_IF;
   IF #statTankLevel < #model.tank.maxLevel THEN #signals.tankSignals.maxLevel := FALSE; END_IF;
END_REGION

REGION Network 11: TANK: recalculate tank level (m³ -> l)
   #signals.tankSignals.actLevel := 1000.0 * #statTankLevel;
END_REGION

REGION Network 12: TANK PRESSURE: calc mass (m = V * p)
   // m = mass [kg]
   // V = volume [m³]
   // p = density [kg/m³]
   #statLiquidMass := #statTankLevel * #model.tank.density;
END_REGION

REGION Network 13: TANK PRESSURE: calc power (F = m * a)
   // F = power [N]
   // m = mass [kg]
   // a = acceleration [m/s²]
   #statLiquidPower := #statLiquidMass * #ACCELERATION;
END_REGION

REGION Network 14: TANK PRESSURE: calc pressure (p = F / A) in [hPa]
   // p = pressure [Pa]
   // F = power [N]
   // A = surface [m²]